      Visibility <- "14_DQ_Data_200CV216ControlOut"
   GraphicView "Graphic view_64" at 581,363 size 107x11; Picture "Graphic_63"
   GraphicView "Graphic view_65" at 695,390 size 12x9; Picture "Graphic_63"
   GraphicView "Graphic view_66" at 851,616 size 24x21; Picture "Graphic_107"
   GraphicView "Graphic view_67" at 1040,616 size 24x21; Picture "Graphic_107"
   IOField "I/O field_8" at 876,617 size 64x18; FormatPattern 99.9; Unit  °C
      ProcessValue <- "12_AI_Data_TIT319_SCALED"
   IOField "I/O field_12" at 1064,617 size 64x18; FormatPattern 99.9; Unit  °C
      ProcessValue <- "12_AI_Data_TIT360_SCALED"
   TextField "Text field_34" at 854,633 size 56x16; Text 'TIT-319'
   TextField "Text field_35" at 1047,633 size 56x16; Text 'TIT-360'
   GraphicView "Graphic view_68" at 1089,539 size 24x21; Picture "Graphic_107"
   TextField "Text field_36" at 1085,559 size 48x16; Text 'LS-001'
   GraphicView "Graphic view_69" at 910,257 size 20x23; Picture "Graphic_36"
   GraphicView "Graphic view_70" at 966,270 size 20x23; Picture "Graphic_36"
   IOField "I/O field_14" at 947,250 size 65x18; FormatPattern s9.99; Unit  bar
      ProcessValue <- "12_AI_Data_PIT316_SCALED"
   GraphicView "Graphic view_71" at 848,241 size 20x26; Picture "Graphic_79"
   TextField "Text field_40" at 433,315 size 70x22; Text 'No Flow'
   TextField "Text field_41" at 433,315 size 70x22; Text '- Flow -'
      Visibility <- "10 DI_DATA_FS115"
      Appearance <- "10 DI_DATA_FS115(1)"
   TextField "Text field_44" at 835,218 size 54x22; Text 'No Flow'
   TextField "Text field_45" at 835,218 size 54x22; Text '- Flow -'
      Visibility <- "10 DI_DATA_FS317"
      Appearance <- "10 DI_DATA_FS317"
   GraphicView "Graphic view_32" at 280,357 size 12x17; Picture "Graphic_64"
   TextField "Text field_48" at 50,404 size 130x20; Text 'I & A Compressor'
      Appearance <- "68_Sys_Status_Data_IA_PRES_IN_RNG"
   GraphicIOField "Graphic I/O field_2" at 273,594 size 196x199; PictureList "IA Compressor_1"
      ProcessValue <- "82_To_HMI_CA Blower Animation"
   GraphicView "Graphic view_13" at 451,640 size 21x27; Picture "Graphic_82"
   GraphicView "Graphic view_36" at 1225,137 size 49x75; Picture "Graphic_108"
   GraphicView "Graphic view_4" at 964,141 size 44x74; Picture "Graphic_108"
   TextField "Text field_50" at 1220,113 size 60x22; Text 'Closed'
      Visibility <- "10_DI_Data_CV401_CLSD"
   IOField "I/O field_5" at 307,295 size 54x22; FormatPattern 999; Unit %
      ProcessValue <- "16_AQ_Data_CV111_CNTRL"
   IOField "I/O field_4" at 307,403 size 54x22; FormatPattern 999; Unit %
      ProcessValue <- "16_AQ_Data_CV203_CNTRL(1)"
   TextField "Text field_52" at 961,125 size 50x16; Text 'CV-403'
   TextField "Text field_53" at 518,576 size 50x16; Text 'CV-127'
   TextField "Text field_56" at 446,576 size 49x16; Text 'PS-101'
   GraphicView "Graphic view_74" at 466,569 size 232x5; Picture "Graphic_63"
   Group "Group_1" at 527,525 size 32x50; Picture "Graphic_72"
   TextField "Text field_54" at 513,526 size 60x22; Text 'Closed'
   TextField "Text field_55" at 513,526 size 60x22; Text 'Opened'
      Visibility <- "14_DQ_Data_200CV127ControlOut"
   GraphicView "Graphic view_73" at 460,550 size 20x26; Picture "Graphic_36"
   GraphicView "Graphic view_75" at 737,434 size 6x141; Picture "Graphic_70"
   GraphicView "Graphic view_78" at 597,569 size 148x5; Picture "Graphic_63"
   GraphicView "Graphic view_3" at 736,566 size 6x8; Picture "Graphic_65"
   GraphicView "Graphic view_28" at 189,356 size 95x11; Picture "Graphic_63"
   GraphicView "Graphic view_19" at 132,317 size 19x12; Picture "Graphic_63"
   GraphicView "Graphic view_72" at 1040,188 size 20x26; Picture "Graphic_36"
   TextField "Text field_59" at 404,73 size 80x18; Text 'Start IGGS'
   TextField "Text field_60" at 340,73 size 70x18; Text 'IA Comp.'
   TextField "Text field_61" at 494,73 size 36x18; Text 'CSW'
   TextField "Text field_62" at 537,73 size 89x18; Text 'Fuel System'
   TextField "Text field_63" at 634,73 size 36x18; Text 'CAB'
   TextField "Text field_64" at 868,72 size 46x18; Text 'Purge'
   TextField "Text field_65" at 806,72 size 52x18; Text 'Pilot B'
   TextField "Text field_66" at 931,72 size 52x18; Text 'Main B'
   TextField "Text field_67" at 1062,72 size 64x18; Text 'Running'
   Circle "Circle_22" at 365,58 size 14x14
      Appearance <- "10 DI_DATA_E131_OK"
   Circle "Circle_23" at 503,58 size 14x14
      Appearance <- "68_Sys_Status_Data_CSW_IL_PRES_IN_RNG"
      Visibility <- "82_To_HMI_IGG RUN Indication"
   Circle "Circle_24" at 572,58 size 14x14
      Visibility <- "68_Sys_Status_Data_CSW_IL_PRES_IN_RNG"
      Appearance <- "68_Sys_Status_Data_FUEL_PRES_IN_RNG(1)"
   Circle "Circle_25" at 642,58 size 14x14
      Visibility <- "68_Sys_Status_Data_FUEL_PRES_IN_RNG(1)"
      Appearance <- "10_DI_Data_E139_RUNNING"
   Circle "Circle_29" at 1080,55 size 20x20
      Appearance <- "14_DQ_Data_24PF1"
   Circle "Circle_31" at 434,58 size 14x14
      Visibility <- "10 DI_DATA_E131_OK"
      Appearance <- "80_From_HMI_RUN_IGG(1)"
   Circle "Circle_32" at 296,58 size 14x14
      Appearance <- "82_To_HMI_CRNT_MODE_IGG"
   Circle "Circle_27" at 822,58 size 14x14
      Visibility <- "102_Pilot_Burner_DB_FLM_DET"
      Appearance <- "102_Pilot_Burner_DB_RUNNING"
   Circle "Circle_28" at 949,58 size 14x14
      Visibility <- "102_Pilot_Burner_DB_FLM_DET"
      Appearance <- "103_Main_Burner_DB_RUNNING"
   Circle "Circle_9" at 887,58 size 14x14
      Visibility <- "102_Pilot_Burner_DB_FLM_DET"
      Appearance <- "104_Pilot_Purge_DB_DN_OK"
   GraphicView "Graphic view_79" at 132,353 size 19x12; Picture "Graphic_63"
   Button "HmiScreenItemData_9" at 2,97 size 184x29; TextOn 'Back'; TextOff 'IGGS Control'
   Button "HmiScreenItemData_4" at 23,192 size 75x51; TextOn 'Back'; TextOff 'Stop'; Authorization "Operate"
      ObjectEnable <- "82_To_HMI_CRNT_MODE_IGG"
      on Release: function_efd93a16("IGG Stop Confirm", 0, 0, -1, -1, 1)
   Circle "Circle_20" at 146,143 size 29x29
      Appearance <- "82_To_HMI_IGG RUN Indication"
   Button "HmiScreenItemData_3" at 23,130 size 75x51; TextOn 'Back'; TextOff 'Start'; Authorization "Operate"
      ObjectEnable <- "82_To_HMI_CRNT_MODE_IGG"
      on Release: function_efd93a16("IGG Start Confirm", 0, 0, -1, -1, 1)
   GraphicView "Graphic view_37" at 684,364 size 11x16; Picture "Graphic_67"
   IOField "I/O field_21" at 635,523 size 80x21; FormatPattern s9999; Unit  mBar
      ProcessValue <- "12_AI_Data_PIT102_SCALED(1)"
   TextField "Text field_68" at 644,576 size 56x16; Text 'PIT-102'
   TextField "Text field_15" at 513,121 size 60x22; Text 'Closed'
   TextField "Text field_16" at 513,121 size 60x22; Text 'Opened'
      Visibility <- "14_DQ_Data_200CV124ControlOut"
   Button "HmiScreenItemData_2" at 1128,64 size 150x43; TextOn 'Back'; TextOff 'IGGS Setup'
      on Release: ActivateScreen("Inert Gas Generator Setup", 0)
   GraphicView "Graphic view_77" at 1,556 size 42x15; Picture "Graphic_20"
   GraphicView "Graphic view_85" at 809,353 size 178x145; Picture "Graphic_132"
      Visibility <- "103_Main_Burner_DB_DN_OK(1)"
   GraphicView "Graphic view_82" at 784,321 size 237x221; Picture "Graphic_130"
      Visibility <- "103_Main_Burner_DB_DN_OK(1)"
   GraphicView "Graphic view_86" at 194,566 size 15x144; Picture "Graphic_101"
   GraphicView "Graphic view_87" at 183,704 size 25x21; Picture "Graphic_97"
   TextField "Text field_69" at 1133,358 size 57x18; Text 'Oxygen'
   IOField "I/O field_22" at 1195,354 size 77x27; FormatPattern 99.99; Unit  %
      ProcessValue <- "12_AI_Data_E600O2ContentIn"
   TextField "Text field_70" at 1150,326 size 121x18; Text 'Inert Gas Profile'
   TextField "Text field_71" at 1133,388 size 67x18; Text 'Setpoint'
   TextField "Text field_72" at 1133,426 size 39x18; Text 'Soot'
   IOField "I/O field_24" at 1195,423 size 77x27; FormatPattern 999.9; Unit  %
      ProcessValue <- "12_AI_Data_E700SootContentIn"
   IOField "I/O field_25" at 1195,460 size 77x27; FormatPattern 999.9; Unit  °C
      ProcessValue <- "12_AI_Data_TIT401_SCALED"
   TextField "Text field_73" at 1133,462 size 47x18; Text 'Temp.'
   IOField "I/O field_26" at 1195,496 size 77x27; FormatPattern 9999; Unit  mBar
      ProcessValue <- "12_AI_Data_PIT402_SCALED"
   TextField "Text field_74" at 1133,500 size 65x18; Text 'Pressure'
   GraphicView "Graphic view_89" at 1116,188 size 20x26; Picture "Graphic_36"
   TextField "Text field_39" at 1097,172 size 59x16; Text 'TIT-401'
   IOField "I/O field_18" at 1095,158 size 63x18; FormatPattern 999.9; Unit  °C
      ProcessValue <- "12_AI_Data_TIT401_SCALED"
   TextField "Text field_46" at 446,526 size 50x22; Text 'P'
      Visibility <- "10 DI_DATA_PS101"
   TextField "Text field_75" at 446,526 size 50x22; Text 'No P'
      Visibility <- "10 DI_DATA_PS101"
      Appearance <- "10 DI_DATA_PS101"
   TextField "Text field_77" at 986,271 size 59x16; Text 'PIT-316'
   TextField "Text field_78" at 882,304 size 56x16; Text 'TIT-315'
   TextField "Text field_79" at 793,221 size 48x16; Text 'FS-317'
   IOField "I/O field_3" at 356,319 size 74x18; FormatPattern s99.99; Unit  Bar
      ProcessValue <- "12_AI_Data_PIT113In_SCALED"
   Button "HmiScreenItemData_7" at 215,117 size 150x43; TextOn 'Back'; TextOff 'Air/Fuel Monitoring'
      on Release: ActivateScreen("Air Fuel Monitoring", 0)
   TextField "Text field_51" at 1220,113 size 60x22; Text 'Opened'
      Visibility <- "10_DI_Data_CV401_OPN"
   Button "HmiScreenItemData_11" at 255,608 size 200x179; TextOn 'Back'; TextOff 'Text'
      on Release: ActivateScreen("Air System", 0)
   Line "Line_4" at 812,352 size 3x22
      Visibility <- "14_DQ_Data_X001ControlOut"
   GraphicView "Graphic view_84" at 796,344 size 38x82; Picture "Graphic_129"
      Visibility <- "102_Pilot_Burner_DB_STATE"
   Button "HmiScreenItemData_13" at 741,647 size 358x51; TextOn 'Back'; TextOff 'Cooling System'
      on Release: ActivateScreen("Cooling System", 0)
   IOField "I/O field_23" at 1195,386 size 77x27; Authorization "User administration"; FormatPattern 99.99; Unit  %
      ProcessValue <- "84_Setpoints_E600_BWT_Target"
   TextField "Text field_91" at 465,759 size 169x20; Text 'Combustion Air Blower'
      Appearance <- "10_DI_Data_E139_VSD_FLT"
   TextField "Text field_88" at 835,190 size 54x22; Text 'No Flow'
   TextField "Text field_92" at 835,190 size 54x22; Text '- Flow -'
      Visibility <- "10 DI_DATA_FS320"
      Appearance <- "10 DI_DATA_FS320"
   TextField "Text field_93" at 793,193 size 48x16; Text 'FS-320'
   Button "HmiScreenItemData_18" at 742,647 size 356x51; TextOn 'Back'; TextOff 'Cooling System'
      on Release: ActivateScreen("Cooling System", 0)
      Visibility <- "51_SLAVE_STATUS_P301_ENBLD"
   IOField "I/O field_33" at 462,699 size 72x25; Authorization "Commissioning"; FormatPattern 9999; Unit  rpm
      ProcessValue <- "80_From_HMI_E139_SET_SPEED"
   IOField "I/O field_34" at 1017,134 size 66x23; FormatPattern 999; Unit  mBar
      ProcessValue <- "19_AUTO_CMNDS_Data_PIT402_Target"
      Appearance <- "19_AUTO_CMNDS_Data_PIT402_Target"
   Button "HmiScreenItemData_19" at 1186,568 size 83x29; TextOn 'Back'; TextOff 'Gas - Trend'
      on Click: function_efd93a16("CV 403 Grafics", 200, 100, -1, -1, 1)
   TextField "Text field_100" at 886,320 size 49x16; Text 'TS-006'
   TextField "Text field_90" at 1117,537 size 54x22; Text 'Text'
   TextField "Text field_38" at 1117,537 size 60x22; Text 'Normal'
      Visibility <- "10 DI_DATA_LS001"
      Appearance <- "10 DI_DATA_LS001"
   TextField "Text field_37" at 1117,537 size 60x22; Text 'Hi Level'
      Visibility <- "10 DI_DATA_LS001"
      Appearance <- "84_Setpoints_TIT315_High"
   GraphicView "Graphic view_90" at 1183,190 size 20x23; Picture "Graphic_36"
   TextField "Text field_103" at 1167,172 size 52x16; Text 'TS-403'
   TextField "Text field_104" at 940,317 size 54x22; Text 'Text'
   TextField "Text field_101" at 940,317 size 54x22; Text 'Hi Temp'
      Visibility <- "10 DI_DATA_TS006(1)"
      Appearance <- "10 DI_DATA_TS006(1)"
   TextField "Text field_102" at 940,317 size 54x22; Text 'Normal'
      Visibility <- "10 DI_DATA_TS006(1)"
   TextField "Text field_107" at 1166,150 size 54x22; Text 'Hi Temp'
      Visibility <- "10 DI_DATA_TS403_FAULT(2)"
      Appearance <- "10 DI_DATA_TS403_FAULT(2)"
   TextField "Text field_108" at 1166,150 size 54x22; Text 'Normal'
      Visibility <- "10 DI_DATA_TS403_FAULT(2)"
      Appearance <- "10 DI_DATA_TS403_FAULT"
   IOField "I/O field_13" at 888,237 size 63x18; FormatPattern 999.9; Unit  °C
      ProcessValue <- "12_AI_Data_TIT315_SCALED"
   IOField "I/O field_20" at 1012,158 size 76x18; FormatPattern s9999; Unit  mBar
      ProcessValue <- "12_AI_Data_PIT402_SCALED"
   GraphicView "Graphic view_88" at 1,713 size 199x13; Picture "Graphic_20"
   TextField "Text field_106" at 886,95 size 59x18; Text 'OPENED'
   GraphicView "Graphic view_1" at 976,199 size 26x62; Picture "Graphic_17"
   TextField "Text field_49" at 1223,246 size 53x16; Text 'CV-401'
   TextField "Text field_76" at 1021,172 size 59x16; Text 'PIT-402'
   GraphicView "Graphic view_60" at 1238,195 size 26x62; Picture "Graphic_17"
   IOField "I/O field_2" at 462,728 size 72x25; FormatPattern 9999; Unit  RPM
      ProcessValue <- "12_AI_Data_E139_RPM_SCALED"
   TextField "Text field_114" at 567,701 size 49x18; Text 'SPEED'
   Button "HmiScreenItemData_15" at 1186,604 size 83x29; TextOn 'Back'; TextOff 'Oxygen'
      on Click: function_efd93a16("CV 203 Grafics", 200, 100, -1, -1, 1)
   IOField "I/O field_28" at 767,752 size 69x23; FormatPattern 999; Unit  mBar
      ProcessValue <- "19_AUTO_CMNDS_Data_PIT402_Target"
      Appearance <- "19_AUTO_CMNDS_Data_PIT402_Target"
   IOField "I/O field_31" at 1034,752 size 80x23; FormatPattern 99.99; Unit  bar
      ProcessValue <- "84_Setpoints_PIT205_Target"
      Appearance <- "84_Setpoints_PIT205_Target"
   TextField "Text field_99" at 1006,724 size 144x20; Text 'Main Fuel Pressure'
   Bar "Bar_1" at 161,270 size 20x105; Unit  %; MinimumValue 0; MaximumValue 100
      ProcessValue <- "12_AI_Data_PIT112In_SCALED"
      MaximumValue <- "84_Setpoints_PIT112_HighHigh"
   TextField "Text field_116" at 52,355 size 57x25; Text 'Enabled'
      Visibility <- "14_DQ_Data_E131ControlOut"
   TextField "Text field_118" at 52,332 size 57x25; Text 'Running'
      Visibility <- "10 DI_DATA_E131_OK"
   IOField "I/O field_17" at 819,414 size 65x25; FormatPattern 999; Unit %
      Visibility <- "10 DI_DATA_FD001_OK"
      ProcessValue <- "12_AI_Data_FD001FlameSignalIn"
   Group "Group_9" at 251,73 size 104x19
   Button "HmiScreenItemData_10" at 14,442 size 178x274; TextOn 'Back'; TextOff 'Text'
      on Release: ActivateScreen("Fuel System", 0)
   DateTimeField "HmiScreenItemData_17" at 1175,0 size 105x30
   DateTimeField "HmiScreenItemData" at 1175,30 size 105x30
   AlarmView "Alarm view_1" at 0,777 size 1280x23
   IOField "I/O field_27" at 744,101 size 83x26; Authorization "Commissioning"; FormatPattern 999; Unit  step
      ProcessValue <- "100_IGG_AUTO_SEQ_DB_CRNT_STEP"
   IOField "I/O field_30" at 744,129 size 83x26; Authorization "Commissioning"; FormatPattern 999; Unit  step
      ProcessValue <- "100_BC_AUTO_SEQ_DB_CRNT_STEP"
   Button "HmiScreenItemData_27" at 633,101 size 83x26; TextOn 'Back'; TextOff 'IGG PLC'
   Button "HmiScreenItemData_28" at 633,129 size 83x26; TextOn 'Back'; TextOff 'BC PLC'
   Group "Group_12" at 677,42 size 115x51
   Circle "Circle_2" at 1013,57 size 14x14
      Visibility <- "102_Pilot_Burner_DB_FLM_DET"
      Appearance <- "19_AUTO_CMNDS_Data_CV203_RAMP_CNTRL"
   TextField "Text field_80" at 984,72 size 82x18; Text 'O2 Control'
   Button "HmiScreenItemData_16" at 209,109 size 376x490; TextOn 'Back'; TextOff 'Text'; Authorization "Operate"
      on Release: ActivateScreen("Air Fuel Monitoring", 0)
   Button "HmiScreenItemData_29" at 770,294 size 329x283; TextOn 'Back'; TextOff 'Text'; Authorization "Commissioning"
      on Release: ActivateScreen("O2 Content Monitoring", 0)
   Button "HmiScreenItemData_30" at 1098,647 size 176x51; TextOn 'FRESH WATER SYSTEM'; TextOff 'Fresh Water System'; Authorization "Operating Mode"
      on Release: ActivateScreen("Fresh Water System", 0)
      Visibility <- "80_From_HMI_P305_PRSNT"
   Button "HmiScreenItemData_31" at 917,134 size 153x117; TextOn 'Back'; TextOff 'Text'
      on Click: function_efd93a16("CV 403 Grafics", 200, 100, -1, -1, 1)
   GraphicView "Graphic view_81" at 662,544 size 20x26; Picture "Graphic_36"
   Group "Group_10" at 434,121 size 70x22
   GraphicView "Graphic view_83" at 1158,203 size 96x48; Picture "Graphic_235"
   Button "HmiScreenItemData_5" at 1165,191 size 114x70; TextOn 'Back'; TextOff 'Text'
      on Press: ActivateScreen("Inert Gas Conditioning Plant", 0)
   Button "HmiScreenItemData_12" at 1117,260 size 158x52; TextOn 'INERT GAS TRANSFER'; TextOff 'Inert Gas Transfer'; TextList "IG Transfer"; Authorization "Operate"
      on Release: ActivateScreen("IG Transfer Mode", 0)
      ProcessValue <- "80_From_HMI_BWT_BYPASS"
   Button "HmiScreenItemData_14" at 1186,533 size 83x29; TextOn 'Back'; TextOff 'Temp-Trends'
      on Click: function_efd93a16("IGG Temperature Trends", 200, 100, -1, -1, 1)
   Button "HmiScreenItemData_20" at 14,127 size 162x117; TextOn 'Back'; TextOff 'Text'
      on Click: function_efd93a16("IGG Control from CCR Warning", 0, 0, 1, -1, 1)
      Visibility <- "user_group"
   Group "Group_13" at 935,209 size 223x226
   Group "Group_14" at 473,288 size 237x372
   Group "Group_15" at 4,254 size 821x468
   Button "HmiScreenItemData_8" at 7,250 size 189x152; TextOn 'Back'; TextOff 'Text'
      on Release: ActivateScreen("Air System", 0)
   Group "Group_16" at 196,173 size 599x224
   Group "Group_11" at 834,364 size 223x284
   GraphicView "Graphic view_24" at 739,597 size 57x58; Picture "Graphic_302"
      Visibility <- "10_DI_Data_IGG_ESTOP_OK"
   Button "HmiScreenItemData_23" at 677,42 size 115x51; TextOn 'Back'; TextOff 'Burner Off'
      Visibility <- "103_Main_Burner_DB_Status"
   Button "HmiScreenItemData_21" at 677,42 size 115x51; TextOn 'Back'; TextOff 'Start Burner'
      Visibility <- "103_Main_Burner_DB_Status"
   Button "HmiScreenItemData_6" at 677,42 size 115x51; TextOn 'Back'; TextOff 'Burner On'
      Visibility <- "103_Main_Burner_DB_Status"
   Button "HmiScreenItemData_22" at 677,42 size 115x51; TextOn 'Back'; TextOff 'Burner Stopped'
      Visibility <- "103_Main_Burner_DB_Status"
   TextField "Text field_42" at 434,121 size 70x22; Text 'No Flow'
   TextField "Text field_43" at 434,121 size 70x22; Text '- Flow -'
      Visibility <- "10 DI_DATA_FS123"
      Appearance <- "10 DI_DATA_FS123"
   Circle "Circle_139" at 1074,338 size 10x10
      Visibility <- "51_SLAVE_STATUS_MAIN_BURNER_ACTV"
      VerticalMovement <- "Main Burner Animation_DB_Animation"
   Circle "Circle_134" at 1013,394 size 10x10
      Visibility <- "51_SLAVE_STATUS_MAIN_BURNER_ACTV"
      DiagonalMovement <- "Main Burner Animation_DB_Animation"
   Circle "Circle_135" at 1036,425 size 10x10
      Visibility <- "51_SLAVE_STATUS_MAIN_BURNER_ACTV"
      DiagonalMovement <- "Main Burner Animation_DB_Animation"
   Circle "Circle_136" at 1041,382 size 10x10
      Visibility <- "51_SLAVE_STATUS_MAIN_BURNER_ACTV"
      DiagonalMovement <- "Main Burner Animation_DB_Animation"
   Circle "Circle_137" at 1080,390 size 10x10
      Visibility <- "51_SLAVE_STATUS_MAIN_BURNER_ACTV"
      DiagonalMovement <- "Main Burner Animation_DB_Animation"
   Circle "Circle_143" at 1073,220 size 16x16
      HorizontalMovement <- "Main Burner Animation_DB_Animation"
      Visibility <- "10_DI_Data_CV401_OPN"
   Circle "Circle_144" at 1142,218 size 16x16
      HorizontalMovement <- "Main Burner Animation_DB_Animation"
      Visibility <- "10_DI_Data_CV401_OPN"
   Circle "Circle_146" at 1068,296 size 16x16
      Visibility <- "51_SLAVE_STATUS_MAIN_BURNER_ACTV"
      VerticalMovement <- "Main Burner Animation_DB_Animation"
   Circle "Circle_147" at 1066,217 size 16x16
      HorizontalMovement <- "Main Burner Animation_DB_Animation"
      Visibility <- "10_DI_Data_CV401_OPN"
   Circle "Circle_148" at 1124,217 size 16x16
      HorizontalMovement <- "Main Burner Animation_DB_Animation"
      Visibility <- "10_DI_Data_CV401_OPN"
   Circle "Circle_149" at 1067,277 size 16x16
      Visibility <- "51_SLAVE_STATUS_MAIN_BURNER_ACTV"
      VerticalMovement <- "Main Burner Animation_DB_Animation"
   Circle "Circle_21" at 1069,258 size 10x10
      Visibility <- "51_SLAVE_STATUS_MAIN_BURNER_ACTV"
      VerticalMovement <- "Main Burner Animation_DB_Animation"
   Circle "Circle_145" at 1014,224 size 10x10
      Visibility <- "51_SLAVE_STATUS_MAIN_BURNER_ACTV"
      HorizontalMovement <- "Main Burner Animation_DB_Animation"
   Circle "Circle_150" at 935,209 size 10x10
      Visibility <- "51_SLAVE_STATUS_MAIN_BURNER_ACTV"
      VerticalMovement <- "Main Burner Animation_DB_Animation"
   Circle "Circle_140" at 954,224 size 10x10
      Visibility <- "51_SLAVE_STATUS_MAIN_BURNER_ACTV"
      DiagonalMovement <- "Main Burner Animation_DB_Animation"
   Circle "Circle_133" at 1072,290 size 10x10
      Visibility <- "51_SLAVE_STATUS_MAIN_BURNER_ACTV"
      VerticalMovement <- "Main Burner Animation_DB_Animation"
   Circle "Circle_138" at 1031,354 size 10x10
      Visibility <- "51_SLAVE_STATUS_MAIN_BURNER_ACTV"
      DiagonalMovement <- "Main Burner Animation_DB_Animation"
   Circle "Circle_142" at 1070,424 size 10x10
      Visibility <- "51_SLAVE_STATUS_MAIN_BURNER_ACTV"
      DiagonalMovement <- "Main Burner Animation_DB_Animation"
   Circle "Circle_127" at 473,646 size 14x14
      Visibility <- "10_DI_Data_E139_RUNNING"
      HorizontalMovement <- "82_To_HMI_CA Blower Animation"
   Circle "Circle_126" at 525,646 size 14x14
      Visibility <- "10_DI_Data_E139_RUNNING"
      HorizontalMovement <- "82_To_HMI_CA Blower Animation"
   Circle "Circle_128" at 612,622 size 14x14
      Visibility <- "10_DI_Data_E139_RUNNING"
      VerticalMovement <- "82_To_HMI_CA Blower Animation"
   Circle "Circle_129" at 612,517 size 14x14
      Visibility <- "10_DI_Data_E139_RUNNING"
      VerticalMovement <- "82_To_HMI_CA Blower Animation"
   Circle "Circle_130" at 612,412 size 14x14
      Visibility <- "10_DI_Data_E139_RUNNING"
      VerticalMovement <- "82_To_HMI_CA Blower Animation"
   Circle "Circle_131" at 639,288 size 14x14
      Visibility <- "10_DI_Data_E139_RUNNING"
      HorizontalMovement <- "82_To_HMI_CA Blower Animation"
   Circle "Circle_132" at 696,288 size 14x14
      Visibility <- "10_DI_Data_E139_RUNNING"
      HorizontalMovement <- "82_To_HMI_CA Blower Animation"
   Circle "Circle_26" at 4,561 size 6x6
      Visibility <- "68_Sys_Status_Data_FUEL_PRES_IN_RNG(1)"
      HorizontalMovement <- "Ful Pump Ani Animation_DB_Animation"
   Circle "Circle_3" at 44,508 size 6x6
      HorizontalMovement <- "IDB_E500A_Animation_Animation"
      Visibility <- "68_Sys_Status_Data_FUEL_PRES_IN_RNG(1)"
   Circle "Circle_17" at 43,608 size 6x6
      HorizontalMovement <- "IDB_E500B_Animation_Animation"
      Visibility <- "68_Sys_Status_Data_FUEL_PRES_IN_RNG(1)"
   Circle "Circle_10" at 137,609 size 6x6
      Visibility <- "10_DI_Data_E500B_ENBLD"
      HorizontalMovement <- "IDB_E500B_Animation_Animation"
   Circle "Circle_7" at 134,507 size 6x6
      HorizontalMovement <- "IDB_E500A_Animation_Animation"
      Visibility <- "10_DI_Data_E500A_ENBLD"
   Circle "Circle_19" at 175,517 size 6x6
      VerticalMovement <- "IDB_E500A_Animation_Animation"
      Visibility <- "10_DI_Data_E500A_ENBLD"
   Circle "Circle_18" at 175,596 size 6x6
      Visibility <- "10_DI_Data_E500B_ENBLD"
      VerticalMovement <- "IDB_E500B_Animation_Animation"
   Circle "Circle_35" at 95,716 size 6x6
      HorizontalMovement <- "Ful Pump Ani Animation_DB_Animation"
      Visibility <- "68_Sys_Status_Data_FUEL_PRES_IN_RNG(1)"
   Circle "Circle_51" at 191,716 size 6x6
      HorizontalMovement <- "Ful Pump Ani Animation_DB_Animation"
      Visibility <- "68_Sys_Status_Data_FUEL_PRES_IN_RNG(1)"
   Circle "Circle_52" at 199,643 size 6x6
      VerticalMovement <- "Ful Pump Ani Animation_DB_Animation"
      Visibility <- "68_Sys_Status_Data_FUEL_PRES_IN_RNG(1)"
   Circle "Circle_53" at 199,579 size 6x6
      VerticalMovement <- "Ful Pump Ani Animation_DB_Animation"
      Visibility <- "68_Sys_Status_Data_FUEL_PRES_IN_RNG(1)"
   Circle "Circle_36" at 202,562 size 6x6
      HorizontalMovement <- "Ful Pump Ani Animation_DB_Animation"
      Visibility <- "68_Sys_Status_Data_FUEL_PRES_IN_RNG(1)"
   Circle "Circle_34" at 296,555 size 6x6
      VerticalMovement <- "Ful Pump Ani Animation_DB_Animation"
      Visibility <- "68_Sys_Status_Data_FUEL_PRES_IN_RNG(1)"
   Circle "Circle_49" at 296,456 size 6x6
      VerticalMovement <- "Ful Pump Ani Animation_DB_Animation"
      Visibility <- "14_DQ_Data_200CV215ControlOut"
   Circle "Circle_37" at 307,471 size 6x6
      HorizontalMovement <- "Ful Pump Ani Animation_DB_Animation"
      Visibility <- "14_DQ_Data_200CV206ControlOut"
   Circle "Circle_38" at 402,470 size 6x6
      HorizontalMovement <- "Ful Pump Ani Animation_DB_Animation"
      Visibility <- "14_DQ_Data_200CV206ControlOut"
   Circle "Circle_39" at 498,469 size 6x6
      HorizontalMovement <- "Ful Pump Ani Animation_DB_Animation"
      Visibility <- "14_DQ_Data_200CV206ControlOut"
   Circle "Circle_40" at 593,470 size 6x6
      HorizontalMovement <- "Ful Pump Ani Animation_DB_Animation"
      Visibility <- "14_DQ_Data_200CV206ControlOut"
   Circle "Circle_43" at 707,462 size 6x6
      VerticalMovement <- "Ful Pump Ani Animation_DB_Animation"
      Visibility <- "14_DQ_Data_200CV207ControlOut"
   Circle "Circle_50" at 297,358 size 6x6
      VerticalMovement <- "Ful Pump Ani Animation_DB_Animation"
      Visibility <- "14_DQ_Data_200CV215ControlOut"
   Circle "Circle_48" at 302,254 size 6x6
      HorizontalMovement <- "Ful Pump Ani Animation_DB_Animation"
      Visibility <- "14_DQ_Data_200CV215ControlOut"
   Circle "Circle_47" at 405,254 size 6x6
      HorizontalMovement <- "Ful Pump Ani Animation_DB_Animation"
      Visibility <- "14_DQ_Data_200CV215ControlOut"
   Circle "Circle_46" at 509,254 size 6x6
      HorizontalMovement <- "Ful Pump Ani Animation_DB_Animation"
      Visibility <- "14_DQ_Data_200CV215ControlOut"
   Circle "Circle_45" at 612,254 size 6x6
      HorizontalMovement <- "Ful Pump Ani Animation_DB_Animation"
      Visibility <- "14_DQ_Data_200CV215ControlOut"
   Circle "Circle_44" at 716,254 size 6x6
      HorizontalMovement <- "Ful Pump Ani Animation_DB_Animation"
      Visibility <- "14_DQ_Data_200CV215ControlOut"
   Circle "Circle_42" at 819,282 size 6x6
      VerticalMovement <- "Ful Pump Ani Animation_DB_Animation"
      Visibility <- "14_DQ_Data_200CV215ControlOut"
   Circle "Circle_74" at 196,359 size 6x6
      HorizontalMovement <- "IDB_E131_Animation_Animation"
      Visibility <- "68_Sys_Status_Data_IA_PRES_IN_RNG"
   Circle "Circle_56" at 280,359 size 6x6
      VerticalMovement <- "IDB_E131_Animation_Animation"
      Visibility <- "10 DI_DATA_FS123"
   Circle "Circle_67" at 282,366 size 6x6
      HorizontalMovement <- "IDB_E131_Animation_Animation"
      Visibility <- "68_Sys_Status_Data_IA_PRES_IN_RNG"
   Circle "Circle_68" at 347,366 size 6x6
      HorizontalMovement <- "IDB_E131_Animation_Animation"
      Visibility <- "10 DI_DATA_FS115"
   Circle "Circle_69" at 407,366 size 6x6
      HorizontalMovement <- "IDB_E131_Animation_Animation"
      Visibility <- "10 DI_DATA_FS115"
   Circle "Circle_70" at 473,366 size 6x6
      HorizontalMovement <- "IDB_E131_Animation_Animation"
      Visibility <- "10 DI_DATA_FS115"
   Circle "Circle_71" at 539,366 size 6x6
      HorizontalMovement <- "IDB_E131_Animation_Animation"
      Visibility <- "10 DI_DATA_FS115"
   Circle "Circle_72" at 606,366 size 6x6
      HorizontalMovement <- "IDB_E131_Animation_Animation"
      Visibility <- "10 DI_DATA_FS115"
   Circle "Circle_73" at 690,391 size 6x6
      HorizontalMovement <- "IDB_E131_Animation_Animation"
      Visibility <- "10 DI_DATA_FS115"
   Circle "Circle_64" at 280,281 size 6x6
      VerticalMovement <- "IDB_E131_Animation_Animation"
      Visibility <- "10 DI_DATA_FS123"
   Circle "Circle_57" at 287,174 size 6x6
      HorizontalMovement <- "IDB_E131_Animation_Animation"
      Visibility <- "10 DI_DATA_FS123"
   Circle "Circle_58" at 370,174 size 6x6
      HorizontalMovement <- "IDB_E131_Animation_Animation"
      Visibility <- "10 DI_DATA_FS123"
   Circle "Circle_59" at 453,174 size 6x6
      HorizontalMovement <- "IDB_E131_Animation_Animation"
      Visibility <- "10 DI_DATA_FS123"
   Circle "Circle_60" at 526,174 size 6x6
      HorizontalMovement <- "IDB_E131_Animation_Animation"
      Visibility <- "10 DI_DATA_FS123"
   Circle "Circle_61" at 619,173 size 6x6
      HorizontalMovement <- "IDB_E131_Animation_Animation"
      Visibility <- "10 DI_DATA_FS123"
   Circle "Circle_62" at 703,174 size 6x6
      HorizontalMovement <- "IDB_E131_Animation_Animation"
      Visibility <- "10 DI_DATA_FS123"
   Circle "Circle_65" at 786,179 size 6x6
      VerticalMovement <- "IDB_E131_Animation_Animation"
      Visibility <- "10 DI_DATA_FS123"
   Circle "Circle_66" at 786,262 size 6x6
      VerticalMovement <- "IDB_E131_Animation_Animation"
      Visibility <- "10 DI_DATA_FS123"
   Circle "Circle_63" at 789,333 size 6x6
      HorizontalMovement <- "IDB_E131_Animation_Animation"
      Visibility <- "10 DI_DATA_FS123"
   Circle "Circle_104" at 1011,436 size 13x13
      DiagonalMovement <- "CSW_Animation_DB_Animation"
      Visibility <- "10 DI_DATA_FS317"
   Circle "Circle_105" at 1029,410 size 13x13
      DiagonalMovement <- "CSW_Animation_DB_Animation"
      Visibility <- "10 DI_DATA_FS317"
   Circle "Circle_100" at 1038,482 size 13x13
      DiagonalMovement <- "CSW_Animation_DB_Animation"
      Visibility <- "10 DI_DATA_FS317"
   Circle "Circle_98" at 1006,471 size 13x13
      DiagonalMovement <- "CSW_Animation_DB_Animation"
      Visibility <- "10 DI_DATA_FS317"
   Circle "Circle_99" at 1044,458 size 13x13
      DiagonalMovement <- "CSW_Animation_DB_Animation"
      Visibility <- "10 DI_DATA_FS317"
   Circle "Circle_107" at 1038,442 size 13x13
      DiagonalMovement <- "CSW_Animation_DB_Animation"
      Visibility <- "10 DI_DATA_FS317"
   Circle "Circle_94" at 1019,364 size 10x10
      DiagonalMovement <- "CSW_Animation_DB_Animation"
      Visibility <- "10 DI_DATA_FS317"
   Circle "Circle_30" at 1018,602 size 8x8
      DiagonalMovement <- "CSW_Animation_DB_Animation"
      Visibility <- "10 DI_DATA_FS317"
   Circle "Circle_97" at 1028,606 size 8x8
      DiagonalMovement <- "CSW_Animation_DB_Animation"
      Visibility <- "10 DI_DATA_FS317"
   Circle "Circle_102" at 834,640 size 8x8
      DiagonalMovement <- "CSW_Animation_DB_Animation"
      Visibility <- "10 DI_DATA_FS317"
   Circle "Circle_108" at 842,556 size 8x8
      DiagonalMovement <- "CSW_Animation_DB_Animation"
      Visibility <- "10 DI_DATA_FS317"
   Circle "Circle_109" at 953,554 size 8x8
      DiagonalMovement <- "CSW_Animation_DB_Animation"
      Visibility <- "10 DI_DATA_FS317"
   Circle "Circle_96" at 962,520 size 8x8
      DiagonalMovement <- "CSW_Animation_DB_Animation"
      Visibility <- "10 DI_DATA_FS317"

screen "Air Fuel Monitoring" 1280x800, template "Template"
   on GenerateScreen: "TitleUpdater"()
   Gauge "Gauge_1" at 441,189 size 184x184; UnitText '%'; CaptionText 'Open'
      ProcessValue <- "16_AQ_Data_CV111_CNTRL"
   TextField "Text field_10" at 118,229 size 176x20; Text 'Atomising Air Pressure'
   Button "Button_9" at 333,227 size 57x25; TextOn 'Enabled'; TextOff 'Text'
   TextField "Text field_17" at 118,266 size 238x20; Text 'I&A Air Pressure Pilot Setpoint'
   Button "Button_11" at 333,263 size 57x25; TextOn 'Enabled'; TextOff 'Text'
   TextField "Text field_20" at 154,155 size 405x26; Text 'Atomising Air Pressure Control (CV-111)'
   TextField "Text field_12" at 117,339 size 110x20; Text 'Valve Position'
   IOField "I/O field_2" at 333,227 size 74x25; FormatPattern 99.99; Unit  bar
      ProcessValue <- "12_AI_Data_PIT113In_SCALED"
   IOField "I/O field_6" at 333,338 size 74x25; FormatPattern 999.99; Unit  %
      ProcessValue <- "16_AQ_Data_CV111_CNTRL"
   Gauge "Gauge_2" at 441,416 size 184x184; UnitText '%'; CaptionText 'Open'
      ProcessValue <- "16_AQ_Data_CV203_CNTRL(1)"
   TextField "Text field_3" at 118,456 size 160x20; Text 'Burner Fuel Pressure'
   Button "Button_3" at 333,454 size 57x25; TextOn 'Enabled'; TextOff 'Text'
   TextField "Text field_4" at 118,493 size 228x20; Text 'Burner Fuel Pressure Setpoint'
   TextField "Text field_5" at 164,383 size 390x26; Text 'Burner Fuel Pressure Control (CV-203)'
   TextField "Text field_6" at 117,547 size 110x20; Text 'Valve Position'
   IOField "I/O field_1" at 333,454 size 74x25; FormatPattern 99.99; Unit  bar
      ProcessValue <- "12_AI_Data_PIT205In_SCALED"
   IOField "I/O field_5" at 333,546 size 74x25; FormatPattern 999.99; Unit  %
      ProcessValue <- "16_AQ_Data_CV203_CNTRL"
   IOField "I/O field_3" at 333,263 size 74x25; Authorization "Commissioning"; FormatPattern 99.99; Unit  bar
      ProcessValue <- "84_Setpoints_PIT113_Pilot_Target"
   TrendView "Trend view_1" at 703,50 size 572x397
   TrendView "Trend view_2" at 703,452 size 572x323
   Button "HmiScreenItemData_3" at 1,1 size 150x43; TextOn 'Back'; TextOff 'Main Index'
      on Release: ActivateScreen("02 Main Index", 0)
   Button "HmiScreenItemData_1" at 1129,1 size 150x43; TextOn 'I&A Compressor Ok'; TextOff 'Back'
      on Release: function_efd93a16()
   IOField "I/O field_31" at 333,492 size 74x23; FormatPattern 99.99; Unit  bar
      ProcessValue <- "84_Setpoints_PIT205_Target"
      Appearance <- "84_Setpoints_PIT205_Target"
   AlarmView "Alarm view_1" at 0,777 size 1280x23
   Button "HmiScreenItemData_4" at 1129,1 size 150x43; TextOn 'I&A Compressor Ok'; TextOff 'Back'
      on Release: function_efd93a16()
   Group "Group_7" at 213,46 size 373x50
   TextField "Text field_1" at 118,303 size 239x20; Text 'I&A Air Pressure Main Setpoint'
   Button "Button_1" at 333,300 size 57x25; TextOn 'Enabled'; TextOff 'Text'
   IOField "I/O field_4" at 333,300 size 74x25; Authorization "Commissioning"; FormatPattern 99.99; Unit  bar
      ProcessValue <- "84_Setpoints_PIT113_Burner_Target"
   Button "HmiScreenItemData_8" at 227,50 size 355x40; TextOn 'Back'; TextOff 'Text'
   TextField "Screen title" at 213,46 size 373x50; Text 'Screen title'

Template "Template_lite" 1280x800
   Button "HmiScreenItemData_12" at 993,4 size 80x35; TextOn 'WARNING'; TextOff 'Warning'
      on Release: ActivateScreen("04 Alarm Log", 0)
      Visibility <- "62_Warning_Data_WRNG_PRSNT"
   Button "HmiScreenItemData_14" at 1080,4 size 80x35; TextOn 'ALARM'; TextOff 'Alarm'
      on Release: ActivateScreen("04 Alarm Log", 0)
      Visibility <- "60_Alarm_Data_ALRM_PRSNT"
   Button "HmiScreenItemData_20" at 906,4 size 80x35; TextOn 'Back'; TextOff 'Lockout'
      on Click: SetBit("80_From_HMI_Reset_Alarms")
      on Press: function_b14e0dd5("80_From_HMI_RST_LOCKOUT", 0)
      Appearance <- "82_To_HMI_E-STOP LATCHED"
   Button "HmiScreenItemData_24" at 810,3 size 64x35; TextOn 'MUTE'; TextOff 'Mute'
      on Press: function_b14e0dd5("80_From_HMI_SLNCE_BZR", 0)
      Appearance <- "80_From_HMI_SLNCE_BZR"
   GraphicView "Graphic view_24" at 876,3 size 29x41; Picture "Graphic_138"
      Visibility <- "Buzzer"
   Circle "Circle_46" at 265,6 size 26x26
      Visibility <- "TRUE"
      Appearance <- "IGG PLC HEART BEAT"
   Circle "Circle_1" at 235,6 size 26x26
      Visibility <- "TRUE"
      Appearance <- "Setpoint Override_DB_Set Pressure"

screen "PGC System" 1280x800, template "Template"
   Button "HmiScreenItemData_1" at -189,1 size 150x43; TextOn 'Back'; TextOff 'Main Index'
      on Release: ActivateScreen("02 Main Index", 0)
   Gauge "Gauge_1" at 454,351 size 184x184; CaptionText 'Pressure'; UnitText 'Bar'
      ProcessValue <- "12_AI_Data_E_400_PT002_SCALED"
      MaximumValue <- "84_Setpoints_E400_PT002_HighHigh"
   TextField "Text field_20" at 187,312 size 324x26; Text 'Process Gas Discharge Pressure'
   TextField "Text field_7" at 221,72 size 326x26; Text 'Process Gas Compressor Control'
   TextField "Text field_10" at 119,405 size 243x20; Text 'Process Gas Discharge Pressure'
   TextField "Text field_17" at 119,464 size 217x20; Text 'Discharge Pressure Setpoint'
   Button "Button_8" at 117,115 size 240x30; TextOn 'TB3 Enabled'; TextOff 'PGC System Not Running OK'
      Visibility <- "10_DI_DATA_E_400_RUN"
   Button "HmiScreenItemData_12" at 141,237 size 69x51; TextOn 'Back'; TextOff 'Reset'; Authorization "Operate"
      on Press: function_b14e0dd5("140_PGC_HRS_RUN_DB_RST", 0)
   IOField "I/O field_10" at 70,236 size 66x25; FormatPattern 9999; Unit  h
      ProcessValue <- "140_PGC_HRS_RUN_DB_SRV_HRS"
   TextField "Text field_22" at 36,238 size 37x20; Text 'Run'
   TextField "Text field_23" at 36,268 size 37x20; Text 'Set'
   TextField "Text field_24" at 79,212 size 100x20; Text 'Service Hour'
   IOField "I/O field_13" at 222,249 size 75x25; FormatPattern 99999; Unit h
      ProcessValue <- "140_PGC_HRS_RUN_DB_HRS"
   IOField "I/O field_14" at 299,249 size 40x25; FormatPattern 99; Unit m
      ProcessValue <- "140_PGC_HRS_RUN_DB_MINS"
   IOField "I/O field_15" at 341,249 size 40x25; FormatPattern 99; Unit s
      ProcessValue <- "140_PGC_HRS_RUN_DB_SECS"
   Button "Button_7" at 654,76 size 57x25; TextOn 'Alarm'; TextOff 'Service'
      Visibility <- "140_PGC_HRS_RUN_DB_SRVC"
      Appearance <- "140_PGC_HRS_RUN_DB_SRVC"
   Button "Button_15" at 187,173 size 57x25; TextOn 'Enabled'; TextOff 'Disabled'
   Button "Button_16" at 341,173 size 64x25; TextOn 'Alarm'; TextOff 'Text'
   TextField "Text field_14" at 44,175 size 115x20; Text 'PG Compressor'
   TextField "Text field_15" at 191,151 size 60x18; Text 'Enabled'
   TextField "Text field_16" at 266,151 size 64x18; Text 'Running'
   TextField "Text field_18" at 343,150 size 78x18; Text 'Shutdown'
   Button "Button_1" at 264,173 size 57x25; TextOn 'Enabled'; TextOff 'Stopped'
   TextField "Text field_32" at 187,173 size 57x25; Text 'Enabled'
      Visibility <- "10_DI_DATA_E_400_SHTDN"
   TextField "Text field_2" at 264,173 size 57x25; Text 'Running'
      Visibility <- "10_DI_DATA_E_400_RUN"
   Button "Button_3" at 341,173 size 64x25; TextOn 'Enabled'; TextOff 'Normal'
   Button "Button_2" at 341,173 size 69x25; TextOn 'Alarm'; TextOff 'Shutdown'
      Visibility <- "10_DI_DATA_E_400_NOK"
      Appearance <- "10_DI_DATA_E_400_NOK"
   Gauge "Gauge_2" at 454,588 size 184x184; UnitText '°C'; CaptionText 'Temperature'
      ProcessValue <- "12_AI_Data_E_400_TE002_SCALED"
      MaximumValue <- "84_Setpoints_E400_TT002_HighHigh"
   TextField "Text field_1" at 187,549 size 365x26; Text 'Process Gas Discharge Temperature'
   TextField "Text field_3" at 119,641 size 178x20; Text 'Discharge Temperature'
   TextField "Text field_4" at 109,699 size 246x20; Text 'Discharge Temperature Setpoint'
   IOField "I/O field_2" at 332,403 size 66x25; FormatPattern 9.99; Unit  Bar
      ProcessValue <- "12_AI_Data_E_400_PT002_SCALED"
   IOField "I/O field_1" at 334,638 size 66x25; FormatPattern 999; Unit  °C
      ProcessValue <- "12_AI_Data_E_400_TE002_SCALED"
   Button "HmiScreenItemData_11" at 3,1 size 150x43; TextOn 'IGG Plant'; TextOff 'GCU Plant'
      on Release: ActivateScreen("Inert Gas Conditioning Plant", 0)
   IOField "I/O field_3" at 332,462 size 66x25; Authorization "Commissioning"; FormatPattern 9.99; Unit  Bar
      ProcessValue <- "84_Setpoints_E400_PT002_HighHigh"
   IOField "I/O field_4" at 334,697 size 66x25; Authorization "Commissioning"; FormatPattern 999; Unit  °C
      ProcessValue <- "84_Setpoints_E400_TT002_HighHigh"
   GraphicView "Graphic view_1" at 514,109 size 192x199; Picture "Graphic_251"
   Button "HmiScreenItemData_3" at 1125,1 size 150x43; TextOn 'I&A Compressor Ok'; TextOff 'Back'
      on Release: function_efd93a16()
   TextField "Text field_5" at 222,226 size 160x25; Text 'Total Run Time'
   TextField "Text field_6" at 818,74 size 312x26; Text 'Process Gas Compressor Purge'
   TextField "Text field_8" at 717,177 size 263x20; Text 'Process Gas Compresor Stop Delay'
   TextField "Text field_11" at 716,111 size 305x20; Text 'Combustion Air Blower after Start Delay'
   IOField "I/O field_7" at 993,109 size 66x25; FormatPattern 999; Unit s
      ProcessValue <- "PGC Flush_DB_CAB after Start Delay"
   TextField "Text field_12" at 716,144 size 208x20; Text 'Combustion Air Blower RPM'
   IOField "I/O field_8" at 993,142 size 66x25; FormatPattern 999; Unit RPM
      ProcessValue <- "PGC Flush_DB_CAB RPM Cmnd"
   Button "HmiScreenItemData_2" at 982,285 size 82x35; TextOn 'Back'; TextOff 'Override'; Authorization "Operating Mode"
      on Press: function_b14e0dd5("PGC Flush_DB_Override", 0)
      Appearance <- "PGC Flush_DB_Flip Flop_Override_Output"
   TextField "Text field_9" at 1068,149 size 91x21; Text 'Running'
      Appearance <- "PGC Flush_DB_Running"
   TextField "Text field_13" at 1068,129 size 91x21; Text 'Enabled'
      Appearance <- "PGC Flush_DB_Activate"
   TextField "Text field_19" at 1068,329 size 91x21; Text 'Done'
      Appearance <- "PGC Flush_DB_Done"
   TextField "Text field_21" at 1068,169 size 91x21; Text 'Open CV405'
      Appearance <- "PGC Flush_DB_CV405 Open"
   TextField "Text field_25" at 1068,189 size 91x21; Text 'Open CV401'
      Appearance <- "PGC Flush_DB_CV401 Open"
   TextField "Text field_26" at 1068,209 size 91x21; Text 'Open CV431'
      Appearance <- "PGC Flush_DB_CV431 Open"
   TextField "Text field_27" at 1068,249 size 91x21; Text 'Close CV441'
      Appearance <- "PGC Flush_DB_CV431 Open"
   TextField "Text field_28" at 1068,269 size 91x21; Text 'Start CAB'
      Appearance <- "PGC Flush_DB_CAB Start"
   TextField "Text field_29" at 1068,289 size 91x21; Text 'Mdlt CV403'
      Appearance <- "PGC Flush_DB_CV403 Modulate"
   TextField "Text field_30" at 1068,309 size 91x21; Text 'Stop PGC'
      Appearance <- "PGC Flush_DB_Stop PGC"
   IOField "I/O field_37" at 890,603 size 90x29; Authorization "Commissioning"; FormatPattern 999; Unit  step
      ProcessValue <- "2110_BTCS_CNTRL_DB_BTCS_STEP"
   Button "HmiScreenItemData_10" at 749,604 size 137x29; TextOn 'Back'; TextOff 'BWTS Step'
   Button "HmiScreenItemData_51" at 749,671 size 137x29; TextOn 'Back'; TextOff 'BWTS State'
   Button "HmiScreenItemData_54" at 749,633 size 495x29; TextOn 'Back'; TextOff 'IGG STEP'; TextList "STEP LIST BTCS"
      ProcessValue <- "2110_BTCS_CNTRL_DB_BTCS_STEP"
   Button "HmiScreenItemData_55" at 749,700 size 495x29; TextOn 'Back'; TextOff 'IGG STEP'; TextList "STATE LIST BTCS"
      ProcessValue <- "2110_BTCS_CNTRL_DB_BTCS_STATE"
   IOField "I/O field_38" at 890,671 size 90x29; Authorization "Commissioning"; FormatPattern 9; Unit  state
      ProcessValue <- "2110_BTCS_CNTRL_DB_BTCS_STATE"
   TextField "Text field_31" at 716,210 size 149x20; Text 'PGC Purge Duration'
   IOField "I/O field_6" at 993,208 size 66x25; FormatPattern 999; Unit m
      ProcessValue <- "PGC Flush_DB_PGC Purge Duration"
   TextField "Text field_33" at 1068,229 size 91x21; Text 'Open CV403'
      Appearance <- "PGC Flush_DB_CV403 Open"
   TextField "Text field_34" at 768,296 size 175x18; Text 'Purge Request Simulate'
      Visibility <- "user_group"
   Switch "Switch_1" at 726,288 size 32x29; CaptionText 'Switch'; TextOn 'ON'; TextOff 'OFF'; Authorization "User administration"; PictureOff "Design_5_PilotLight_Green_Off"; PictureOn "Design_5_PilotLight_Green_On"
      on Change: InvertBit("Sequence Times_DB_Treatment Timer_Enable")
      Visibility <- "user_group"
      ProcessValue <- "19_AUTO_CMNDS_Data_Purge Rqst Simulate"
   TextField "Text field_35" at 1160,149 size 106x21; Text 'Running'
      Appearance <- "PGC Flush_DB_Running"
   TextField "Text field_36" at 1160,129 size 106x21; Text 'Enabled'
      Appearance <- "PGC Flush_DB_Activate"
   TextField "Text field_37" at 1160,329 size 106x21; Text 'Done'
      Appearance <- "100_GCU_AUTO_SEQ_DB_CRNT_STEP"
   TextField "Text field_38" at 1160,169 size 106x21; Text 'Opened CV405'
      Appearance <- "1405_PID_CV405_ManualEnable"
   TextField "Text field_39" at 1160,189 size 106x21; Text 'Opened CV401'
      Appearance <- "PGC Flush_DB_CV401 Opened"
   TextField "Text field_40" at 1160,209 size 106x21; Text 'Opened CV431'
      Appearance <- "PGC Flush_DB_CV431 Opened"
   TextField "Text field_41" at 1160,249 size 106x21; Text 'Closed CV441'
      Appearance <- "PGC Flush_DB_CV441 Closed"
   TextField "Text field_42" at 1160,269 size 106x21; Text 'Started CAB'
      Appearance <- "PGC Flush_DB_CAB Started"
   TextField "Text field_43" at 1160,289 size 106x21; Text 'Mdling CV403'
      Appearance <- "1403_PID_300CV403_ModeActivate"
   TextField "Text field_44" at 1160,309 size 106x21; Text 'Stoped PGC'
      Appearance <- "PGC Flush_DB_PGC Stoped"
   TextField "Text field_45" at 1160,229 size 106x21; Text 'Opened CV403'
      Appearance <- "1403_PID_300CV403_ManualEnable"
   TextField "Text field_46" at 711,332 size 173x20; Text 'Air / Inert Gas Pressure'
   Button "Button_9" at 1001,329 size 57x25; TextOn 'Enabled'; TextOff 'Text'
   TextField "Text field_47" at 710,366 size 277x20; Text 'Air / Inert Gas Pressure Setpoint (Pre-Ignition)'
   Button "Button_11" at 1001,364 size 57x25; TextOn 'Enabled'; TextOff 'Text'
   TextField "Text field_48" at 718,498 size 182x20; Text 'Modulating Valve Position'
   TextField "Text field_49" at 709,399 size 278x20; Text 'Air / Inert Gas Pressure Setpoint (Main-Ignition)'
   Button "Button_10" at 1001,397 size 57x25; TextOn 'Enabled'; TextOff 'Text'
   IOField "I/O field_9" at 993,329 size 66x25; FormatPattern 999; Unit  mbar
      ProcessValue <- "12_AI_Data_PIT402_SCALED"
   IOField "I/O field_12" at 993,364 size 66x25; Authorization "Commissioning"; FormatPattern 999; Unit  mbar
      ProcessValue <- "84_Setpoints_PIT402_Pilot_Target"
   IOField "I/O field_16" at 993,495 size 66x25; FormatPattern 999; Unit  %
      ProcessValue <- "16_AQ_Data_CV403_CNTRL"
   IOField "I/O field_17" at 993,462 size 66x25; FormatPattern 999; Unit  mBar
      ProcessValue <- "19_AUTO_CMNDS_Data_PIT402_Target"
      Appearance <- "19_AUTO_CMNDS_Data_PIT402_Target"
   IOField "I/O field_18" at 993,396 size 66x25; Authorization "Commissioning"; FormatPattern 999; Unit  mbar
      ProcessValue <- "84_Setpoints_PIT402_Main_Target"
   TextField "Text field_50" at 1068,497 size 58x20; Text 'Opened'
   TextField "Text field_51" at 711,465 size 266x20; Text 'Air / Inert Gas Pressure Setpoint (Current)'
   TextField "Text field_52" at 709,432 size 278x20; Text 'Air / Inert Gas Pressure Setpoint (Post-Ignition)'
   Button "Button_4" at 1001,430 size 57x25; TextOn 'Enabled'; TextOff 'Text'
   IOField "I/O field_19" at 993,429 size 66x25; Authorization "Commissioning"; FormatPattern 999; Unit  mbar
      ProcessValue <- "84_Setpoints_PIT401_Post_Target_Max"
   TextField "Text field_53" at 1079,107 size 73x20; Text 'Command'
   TextField "Text field_54" at 1182,107 size 73x20; Text 'Feedback'
   IOField "I/O field_20" at 70,266 size 66x25; Authorization "Commissioning"; FormatPattern 9999; Unit h
      ProcessValue <- "140_PGC_HRS_RUN_DB_SHRS_IP"
   TextField "Text field_55" at 716,243 size 168x20; Text 'Temperature Setpoint'
   IOField "I/O field_11" at 993,241 size 66x25; FormatPattern 999; Unit  °C
      ProcessValue <- "PGC Flush_DB_Temperature Setpoint"
   Button "HmiScreenItemData_19" at 749,567 size 495x29; TextOn 'Back'; TextOff 'IGG STEP'; TextList "STEP LIST_GCU"
      ProcessValue <- "100_GCU_AUTO_SEQ_DB_CRNT_STEP"
   IOField "I/O field_21" at 890,537 size 90x29; Authorization "Commissioning"; FormatPattern 999; Unit  Step
      ProcessValue <- "100_GCU_AUTO_SEQ_DB_CRNT_STEP"
   Button "HmiScreenItemData_9" at 749,536 size 100x30; TextOn 'Back'; TextOff 'GCU PLC'
   Button "HmiScreenItemData_16" at 238,742 size 83x29; TextOn 'Back'; TextOff 'Temp-Trends'
      on Click: function_efd93a16("PGC Temperature Trends", 200, 100, -1, -1, 1)
   IOField "I/O field_22" at 993,175 size 66x25; FormatPattern 999; Unit m
      ProcessValue <- "PGC Flush_DB_PGC Stop Delay"

